        [16].12   // Node 3 message write error flag
        [0].12   // Node 2 Message Write Error Flag
        [32].12   // Node 4 message write error flag
        [48].12   // Node 5 message write error flag
        [64].12   // Node 6 message write error flag
        [16]   // Node 3 message write output data control block
        [80].12   // Node 7 message write error flag
        [96].12   // Node 8 message write error flag
        [2]   // FV2 Temperature Scaled -100/+400 tenths degree C
   FV_N101 : INT[255] := ([0] := 152, [1] := 60, [2] := 60, [3] := 586, [4] := 32767, [5] := 1107, [6] := 169, [7] := 117, [9] := 70, [10] := 110);   // FV INT Fermentation control integer workspace
        [9]   // Temp.register
        [7]   // Pointer to vessel's data file
        [35]   // Checkword Pointer
        [0]   // FV Data File Pointer
        [4]   // Next breakpoint time
        [1]   // Setpoint at previous breakpoint
        [30]   // PV550 Manual Valve Control Valve Checkword Number
        [2]   // Setpoint at next breakpoint
        [12]   // Operator Interface CT1 Manual Operation Value
        [14]   // Operator Interface CT2 Manual Operation Value
        [3]   // Previous breakpoint time
        [16]   // Operator Interface CT3 Manual Operation Value
        [18]   // Operator Interface CT4 Manual Operation Value
        [30].15   // Stops Invalid Pointer Error If No Valves Selected On Op. Int
        [20]   // Operator Interface CT5 Manual Operation Value
        [22]   // Operator Interface CT6 Manual Operation Value
        [38]   // Copy Of Current Checkword Manual Enabled Flag
        [32]   // Copy Of Current Checkword Energised Input Flag
        [37]   // Copy Of Current Checkword Energised Input Flag
        [36]   // Valve Operation 1 Open 2 Close 3 Auto
        [8]   // Fermenting Room PV550 data file pointer
        [6]   // Temporary result register
        [15].0   // Current Valve Manual/ Auto(PLC)
        [11].0   // Current Valve Energised/ De-energised
        [13].0   // Current Valve Energised/ De-energised
        [5]   // Time since last B.P in 1/10 hour
   FV_N104 : INT[255] := ([0] := -32768, [1] := -32768, [2] := -32768, [3] := -32768, [4] := -32768, [5] := -32768, [6] := -32768, [7] := -32768, [8] := -32768, [9] := -32768, [10] := -32768, [11] := -32768, [12] := -32768, [13] := -32768, [14] := -32768, [15] := -32768, [16] := -32768, [17] := -32768, [18] := -32768, [19] := -32768, [20] := -32768, [21] := -32768, [22] := -32768, [23] := -32768, [24] := -32768);   // FV_PC_BUF PC>PLC Fermentation Control Command Buff er File
        [23]   // PC>PLC FV System Command Buffer Command Type 1=Start,2=Stop 3=Modify Control
        [11]   // PC>PLC FV System Command Buffer Breakpoint F Time
        [13]   // PC>PLC FV System Command Buffer Breakpoint G Time
        [1]   // PC>PLC FV System Command Buffer Breakpoint A Time
        [3]   // PC>PLC FV System Command Buffer Breakpoint B Time
        [5]   // PC>PLC FV System Command Buffer Breakpoint C Time
        [7]   // PC>PLC FV System Command Buffer Breakpoint D Time
        [9]   // PC>PLC FV System Command Buffer Breakpoint E Time
        [2]   // PC>PLC FV System Command Buffer Breakpoint A Temperature Setpoint
        [4]   // PC>PLC FV System Command Buffer Breakpoint B Temperature Setpoint
        [6]   // PC>PLC FV System Command Buffer Breakpoint C Temperature Setpoint
        [8]   // PC>PLC FV System Command Buffer Breakpoint D Temperature Setpoint
        [0]   // PC>PLC FV System Vessel Number 1-28 = FV1-25,YSV1-3 95-96 YST1-2
        [15].4   // FV System PC Command Buffer Control Flags 1=Ageing Profile
        [15].6   // FV System PC Command Buffer Control Flags 1=Wait for yeast
        [10]   // PC>PLC FV System Command Buffer Breakpoint E Temperature Setpoint
        [12]   // PC>PLC FV System Command Buffer Breakpoint F Temperature Setpoint
        [14]   // PC>PLC FV System Command Buffer Breakpoint G Temperature Setpoint
        [15]   // PC>PLC FV System Command Buffer Profile Control / Configuration Flags
        [24]   // FV System PC Command Buffer Phase Number
        [16]   // PC>PLC FV System Command Buffer PC Private Flags
   FV_N11 : INT[255] := ([0] := 1, [32] := -1028);   // LOOP NO.
        [11].0   // Me>Node 5 heartbeat bit
        [14].0   // Me>Node 6 heartbeat bit
        [17].0   // Me>Node 7 heartbeat bit
        [20].0   // Me>Node 8 heartbeat bit
        [9].1   // BHP_RS Borehole Pump Start Signal Node 5 Output 1
        [2]   // Me>Node 2 Flags
        [0].0   // NODE 2 Outputs CT1 cooling valve drive flag
        [0]   // Check Loop Counter In Range
        [0].1   // NODE 2 Outputs CT2 cooling valve drive flag
        [11].1   // Node 5 to resend data
        [14].1   // Node 6 to resend data
        [0].6   // NODE 2 Outputs Fridge 1 Remote Start flag
        [0].2   // NODE 2 Outputs CT3 cooling valve drive flag
        [0].3   // NODE 2 Outputs CT4 cooling valve drive flag
        [170]   // Me>Node 7 heartbeat bit
        [17].1   // Node 7 to resend data
        [20].1   // Node 8 to resend data
        [2].0   // Me>Node 2 heartbeat bit
        [0].7   // NODE 2 Outputs Glycol recirc pump start flag
        [5].0   // Me>Node 3 heartbeat bit
        [0].4   // NODE 2 Outputs CT5 cooling valve drive flag
        [8].0   // Me>Node 4 heartbeat bit
        [0].5   // NODE 2 Outputs CT6 cooling valve drive flag
        [15]   // Move Binary Image Back To Node 7 Outputs
        [2].1   // Node 2 to resend data
        [5].1   // Node 3 to resend data
        [8].1   // Node 4 to resend data
   FV_N110 : INT[255] := ([0] := 231, [2] := 170, [3] := 100, [4] := 190, [5] := 275, [6] := 190, [7] := 305, [8] := 160, [9] := 486, [10] := 160, [11] := 586, [12] := 60, [13] := 32767, [14] := 60, [15] := 64, [17] := -32767, [18] := -32767, [19] := 1680, [20] := 13, [22] := 1693, [23] := 3, [24] := 6, [25] := 60, [26] := 60, [27] := 1693, [29] := 2, [30] := 24, [40] := 3, [41] := 59);   // FV DATA 0 CURRENT FV DATA
        [29]   // FLAGS - PLC CONTROL
        [28]   // CURRENT VOLUME HL*10
        [41]   // Cone ACTUAL TEMPERATURE -DEGREES 'C'*10
        [19]   // Current FV max. fermentation time
        [1]   // TEMPERATURE BREAKPOINT A. TIME 1/10 HOURS(ALWAYS=0)
        [29].1   // Current vessel deferred chilling enabled flag
        [3]   // TEMPERATURE BREAKPOINT B. TIME 1/10 HOURS(ALWAYS=0)
        [11]   // TEMPERATURE BREAKPOINT F. TIME 1/10 HOURS(ALWAYS=0)
        [13]   // TEMPERATURE BREAKPOINT G. TIME 1/10 HOURS(ALWAYS=0)
        [5]   // TEMPERATURE BREAKPOINT C. TIME 1/10 HOURS(ALWAYS=0)
        [7]   // TEMPERATURE BREAKPOINT D. TIME 1/10 HOURS(ALWAYS=0)
        [9]   // TEMPERATURE BREAKPOINT E. TIME 1/10 HOURS(ALWAYS=0)
        [30].5   // Current vessel deferred chilling temp.high flag
        [22]   // Current FV total residence time
        [15].5   // Profile Control Flags : This is a conditioning profile
        [15].3   // PLC TO USE CONE COOLING JACKET
        [15].9   // Current vessel deferred chilling manual override
        [20]   // Current FV warm conditioning time
        [27]   // CURRENT ELAPSED HOURS *10
        [40]   // FV Routing Status 9=Dirty
        [30].0   // Jacket Cooling Valve to open
        [26]   // Calculated Setpoint 1/10 degrees C
        [29].0   // PC TO SAVE TEMPERATURE DATA
        [15]   // FLAGS-PROFILE CONTROL
        [24]   // Phase0=No control 1to6 =Fermenting 8 =Pitching Hold 10 =Maturation 11to16=Conditioning
        [10]   // TEMPERATURE SETPOINT E. 1/10 DEGREE 'C'
        [15].2   // PLC TO FOLLOW RAMP Breakpoints A to B
        [12]   // TEMPERATURE SETPOINT F. 1/10 DEGREE 'C'
        [14]   // TEMPERATURE SETPOINT G. 1/10 DEGREE 'C'
        [36]   // Current vessel time to deferred chlling start (hrs.x10)
        [16].1   // Profile control flag Hold at B.P B
        [16].2   // Profile control flag Hold at B.P C
        [30].3   // Current vessel deferred chilling active
        [16].3   // Profile control flag Hold at B.P D
        [16].4   // Profile control flag Hold at B.P E
        [0]   // FV SYSTEM WORKING BUFFER VESSEL NUMBER
        [2]   // TEMPERATURE SETPOINT A. 1/10 DEGREE 'C'
        [16].5   // Profile control flag Hold at B.P F
        [16].6   // Profile control flag Hold at B.P G
        [30].4   // Current vessel final temp.reached
        [4]   // TEMPERATURE SETPOINT B. 1/10 DEGREE 'C'
        [6]   // TEMPERATURE SETPOINT C. 1/10 DEGREE 'C'
        [8]   // TEMPERATURE SETPOINT D. 1/10 DEGREE 'C'
        [30].1   // Cone Cooling Valve to open
        [25]   // Jacket ACTUAL TEMPERATURE -DEGREES 'C'*10
        [15].4   // Profile Control Flags : This is a maturation profile
   FV_N111 : INT[50] := ([0] := 1, [2] := 175, [3] := 200, [4] := 200, [5] := 440, [6] := 200, [7] := 480, [8] := 180, [9] := 650, [10] := 180, [11] := 820, [12] := 60, [13] := 32767, [14] := 60, [15] := 64, [16] := 20, [17] := -32767, [18] := -32767, [19] := 1680, [22] := 253, [23] := 1, [24] := 2, [25] := 199, [26] := 200, [27] := 253);   // FV1, CURRENT FV DATA
        [27]   // FV1,CURRENT ELAPSED HOURS *10
        [40]   // FV1,FV Routing Status 9=Dirty
        [36]   // FV1,Current vessel time to deferred chlling start (hrs.x10)
        [30].1   // FV1,Cone Cooling Valve to open
        [15].5   // FV1,Profile Control Flags : This is a conditioning profile
        [15]   // FV1,FLAGS-PROFILE CONTROL
        [30].3   // FV1,Current vessel deferred chilling active
        [24]   // FV1,Phase0=No control 1to6 =Fermenting 8 =Pitching Hold 10 =Maturation 11to16=Conditioning
        [15].4   // FV1,Profile Control Flags : This is a maturation profile
        [25]   // FV1,Jacket ACTUAL TEMPERATURE -DEGREES 'C'*10
        [15].2   // FV1,PLC TO FOLLOW RAMP Breakpoints A to B
        [29]   // FV1,FLAGS - PLC CONTROL
        [0]   // FV1,FV SYSTEM WORKING BUFFER VESSEL NUMBER
        [2]   // FV1,TEMPERATURE SETPOINT A. 1/10 DEGREE 'C'
        [30].4   // FV1,Current vessel final temp.reached
        [4]   // FV1,TEMPERATURE SETPOINT B. 1/10 DEGREE 'C'
        [6]   // FV1,TEMPERATURE SETPOINT C. 1/10 DEGREE 'C'
        [8]   // FV1,TEMPERATURE SETPOINT D. 1/10 DEGREE 'C'
        [11]   // FV1,TEMPERATURE BREAKPOINT F. TIME 1/10 HOURS(ALWAYS=0)
        [13]   // FV1,TEMPERATURE BREAKPOINT G. TIME 1/10 HOURS(ALWAYS=0)
        [30].5   // FV1,Current vessel deferred chilling temp.high flag
        [28]   // FV1,CURRENT VOLUME HL*10
        [15].3   // FV1,PLC TO USE CONE COOLING JACKET
        [41]   // FV1,Cone ACTUAL TEMPERATURE -DEGREES 'C'*10
        [26]   // FV1,Calculated Setpoint 1/10 degrees C
        [19]   // FV1,Current FV max. fermentation time
        [20]   // FV1,Current FV warm conditioning time
        [22]   // FV1,Current FV total residence time
        [29].0   // FV1,PC TO SAVE TEMPERATURE DATA
        [1]   // FV1,TEMPERATURE BREAKPOINT A. TIME 1/10 HOURS(ALWAYS=0)
        [29].1   // FV1,Current vessel deferred chilling enabled flag
        [30].0   // FV1,Jacket Cooling Valve to open
        [3]   // FV1,TEMPERATURE BREAKPOINT B. TIME 1/10 HOURS(ALWAYS=0)
        [5]   // FV1,TEMPERATURE BREAKPOINT C. TIME 1/10 HOURS(ALWAYS=0)
        [7]   // FV1,TEMPERATURE BREAKPOINT D. TIME 1/10 HOURS(ALWAYS=0)
        [9]   // FV1,TEMPERATURE BREAKPOINT E. TIME 1/10 HOURS(ALWAYS=0)
        [16].1   // FV1,Profile control flag Hold at B.P B
        [16].2   // FV1,Profile control flag Hold at B.P C
        [16].3   // FV1,Profile control flag Hold at B.P D
        [16].4   // FV1,Profile control flag Hold at B.P E
        [16].5   // FV1,Profile control flag Hold at B.P F
        [16].6   // FV1,Profile control flag Hold at B.P G
        [10]   // FV1,TEMPERATURE SETPOINT E. 1/10 DEGREE 'C'
        [15].9   // FV1,Current vessel deferred chilling manual override
        [12]   // FV1,TEMPERATURE SETPOINT F. 1/10 DEGREE 'C'
        [14]   // FV1,TEMPERATURE SETPOINT G. 1/10 DEGREE 'C'
   FV_N112 : INT[50] := ([0] := 2, [2] := 170, [3] := 100, [4] := 190, [5] := 264, [6] := 190, [7] := 290, [8] := 160, [9] := 532, [10] := 160, [11] := 632, [12] := 60, [13] := 32767, [14] := 60, [15] := 64, [17] := -32767, [18] := -32767, [19] := 1680, [20] := 15, [22] := 1695, [23] := 3, [24] := 6, [25] := 60, [26] := 60, [27] := 1695, [29] := 2, [30] := 24);   // FV2, CURRENT FV DATA
        [27]   // FV2,CURRENT ELAPSED HOURS *10
        [40]   // FV2,FV Routing Status 9=Dirty
        [36]   // FV2,Current vessel time to deferred chlling start (hrs.x10)
        [30].1   // FV2,Cone Cooling Valve to open
        [15]   // FV2,FLAGS-PROFILE CONTROL
        [15].5   // FV2,Profile Control Flags : This is a conditioning profile
        [30].3   // FV2,Current vessel deferred chilling active
        [24]   // FV2,Phase0=No control 1to6 =Fermenting 8 =Pitching Hold 10 =Maturation 11to16=Conditioning
        [15].4   // FV2,Profile Control Flags : This is a maturation profile
        [25]   // FV2,Jacket ACTUAL TEMPERATURE -DEGREES 'C'*10
        [15].2   // FV2,PLC TO FOLLOW RAMP Breakpoints A to B
        [29]   // FV2,FLAGS - PLC CONTROL
        [0]   // FV2,FV SYSTEM WORKING BUFFER VESSEL NUMBER
        [2]   // FV2,TEMPERATURE SETPOINT A. 1/10 DEGREE 'C'
        [30].4   // FV2,Current vessel final temp.reached
        [4]   // FV2,TEMPERATURE SETPOINT B. 1/10 DEGREE 'C'
        [6]   // FV2,TEMPERATURE SETPOINT C. 1/10 DEGREE 'C'
        [8]   // FV2,TEMPERATURE SETPOINT D. 1/10 DEGREE 'C'
        [11]   // FV2,TEMPERATURE BREAKPOINT F. TIME 1/10 HOURS(ALWAYS=0)
        [13]   // FV2,TEMPERATURE BREAKPOINT G. TIME 1/10 HOURS(ALWAYS=0)
        [15].3   // FV2,PLC TO USE CONE COOLING JACKET
        [30].5   // FV2,Current vessel deferred chilling temp.high flag
        [19]   // FV2,Current FV max. fermentation time
        [28]   // FV2,CURRENT VOLUME HL*10
        [41]   // FV2,Cone ACTUAL TEMPERATURE -DEGREES 'C'*10
        [26]   // FV2,Calculated Setpoint 1/10 degrees C
        [1]   // FV2,TEMPERATURE BREAKPOINT A. TIME 1/10 HOURS(ALWAYS=0)
        [29].1   // FV2,Current vessel deferred chilling enabled flag
        [20]   // FV2,Current FV warm conditioning time
        [3]   // FV2,TEMPERATURE BREAKPOINT B. TIME 1/10 HOURS(ALWAYS=0)
        [22]   // FV2,Current FV total residence time
        [29].0   // FV2,PC TO SAVE TEMPERATURE DATA
        [5]   // FV2,TEMPERATURE BREAKPOINT C. TIME 1/10 HOURS(ALWAYS=0)
        [7]   // FV2,TEMPERATURE BREAKPOINT D. TIME 1/10 HOURS(ALWAYS=0)
        [9]   // FV2,TEMPERATURE BREAKPOINT E. TIME 1/10 HOURS(ALWAYS=0)
        [30].0   // FV2,Jacket Cooling Valve to open
        [16].1   // FV2,Profile control flag Hold at B.P B
        [16].2   // FV2,Profile control flag Hold at B.P C
        [16].3   // FV2,Profile control flag Hold at B.P D
        [16].4   // FV2,Profile control flag Hold at B.P E
        [16].5   // FV2,Profile control flag Hold at B.P F
        [16].6   // FV2,Profile control flag Hold at B.P G
        [15].9   // FV2,Current vessel deferred chilling manual override
        [10]   // FV2,TEMPERATURE SETPOINT E. 1/10 DEGREE 'C'
        [12]   // FV2,TEMPERATURE SETPOINT F. 1/10 DEGREE 'C'
        [14]   // FV2,TEMPERATURE SETPOINT G. 1/10 DEGREE 'C'
   FV_N113 : INT[50] := ([0] := 3, [1] := -32767, [2] := -32767, [3] := -32767, [4] := -32767, [5] := -32767, [6] := -32767, [7] := -32767, [8] := -32767, [9] := -32767, [10] := -32767, [11] := -32767, [12] := -32767, [13] := -32767, [14] := -32767, [15] := -32767, [16] := -32767, [17] := -32767, [18] := -32767, [19] := -32767, [20] := -32767, [21] := -32767, [22] := -32767, [23] := 2, [25] := 431, [30] := 32);   // FV3, CURRENT FV DATA
        [27]   // FV3,CURRENT ELAPSED HOURS *10
        [40]   // FV3,FV Routing Status 9=Dirty
        [36]   // FV3,Current vessel time to deferred chlling start (hrs.x10)
        [30].1   // FV3,Cone Cooling Valve to open
        [15]   // FV3,FLAGS-PROFILE CONTROL
        [15].5   // FV3,Profile Control Flags : This is a conditioning profile
        [30].3   // FV3,Current vessel deferred chilling active
        [24]   // FV3,Phase0=No control 1to6 =Fermenting 8 =Pitching Hold 10 =Maturation 11to16=Conditioning
        [15].4   // FV3,Profile Control Flags : This is a maturation profile
        [25]   // FV3,Jacket ACTUAL TEMPERATURE -DEGREES 'C'*10
        [15].2   // FV3,PLC TO FOLLOW RAMP Breakpoints A to B
        [29]   // FV3,FLAGS - PLC CONTROL
        [0]   // FV3,FV SYSTEM WORKING BUFFER VESSEL NUMBER
        [2]   // FV3,TEMPERATURE SETPOINT A. 1/10 DEGREE 'C'
        [30].4   // FV3,Current vessel final temp.reached
        [4]   // FV3,TEMPERATURE SETPOINT B. 1/10 DEGREE 'C'
        [6]   // FV3,TEMPERATURE SETPOINT C. 1/10 DEGREE 'C'
        [8]   // FV3,TEMPERATURE SETPOINT D. 1/10 DEGREE 'C'
        [19]   // FV3,Current FV max. fermentation time
        [1]   // FV3,TEMPERATURE BREAKPOINT A. TIME 1/10 HOURS(ALWAYS=0)
        [20]   // FV3,Current FV warm conditioning time
        [29].1   // FV3,Current vessel deferred chilling enabled flag
        [3]   // FV3,TEMPERATURE BREAKPOINT B. TIME 1/10 HOURS(ALWAYS=0)
        [11]   // FV3,TEMPERATURE BREAKPOINT F. TIME 1/10 HOURS(ALWAYS=0)
        [13]   // FV3,TEMPERATURE BREAKPOINT G. TIME 1/10 HOURS(ALWAYS=0)
        [30].5   // FV3,Current vessel deferred chilling temp.high flag
        [28]   // FV3,CURRENT VOLUME HL*10
        [5]   // FV3,TEMPERATURE BREAKPOINT C. TIME 1/10 HOURS(ALWAYS=0)
        [15].3   // FV3,PLC TO USE CONE COOLING JACKET
        [26]   // FV3,Calculated Setpoint 1/10 degrees C
        [7]   // FV3,TEMPERATURE BREAKPOINT D. TIME 1/10 HOURS(ALWAYS=0)
        [41]   // FV3,Cone ACTUAL TEMPERATURE -DEGREES 'C'*10
        [9]   // FV3,TEMPERATURE BREAKPOINT E. TIME 1/10 HOURS(ALWAYS=0)
        [22]   // FV3,Current FV total residence time
        [29].0   // FV3,PC TO SAVE TEMPERATURE DATA
        [30].0   // FV3,Jacket Cooling Valve to open
        [16].1   // FV3,Profile control flag Hold at B.P B
        [16].2   // FV3,Profile control flag Hold at B.P C
        [16].3   // FV3,Profile control flag Hold at B.P D
        [10]   // FV3,TEMPERATURE SETPOINT E. 1/10 DEGREE 'C'
        [16].4   // FV3,Profile control flag Hold at B.P E
        [16].5   // FV3,Profile control flag Hold at B.P F
        [16].6   // FV3,Profile control flag Hold at B.P G
        [15].9   // FV3,Current vessel deferred chilling manual override
        [12]   // FV3,TEMPERATURE SETPOINT F. 1/10 DEGREE 'C'
        [14]   // FV3,TEMPERATURE SETPOINT G. 1/10 DEGREE 'C'
   FV_N114 : INT[50] := ([0] := 4, [2] := 240, [3] := 100, [4] := 240, [5] := 280, [6] := 240, [7] := 340, [8] := 240, [9] := 500, [10] := 240, [11] := 710, [12] := 240, [13] := 32767, [14] := 235, [17] := -32767, [18] := -32767, [19] := 14400, [20] := 18367, [22] := 32767, [23] := 3, [24] := 1, [25] := 247, [26] := 240, [27] := -9629, [29] := 2, [30] := 24);   // FV4, CURRENT FV DATA
        [15]   // FV4,FLAGS-PROFILE CONTROL
        [27]   // FV4,CURRENT ELAPSED HOURS *10
        [40]   // FV4,FV Routing Status 9=Dirty
        [36]   // FV4,Current vessel time to deferred chlling start (hrs.x10)
        [30].1   // FV4,Cone Cooling Valve to open
        [15].5   // FV4,Profile Control Flags : This is a conditioning profile
        [30].3   // FV4,Current vessel deferred chilling active
        [24]   // FV4,Phase0=No control 1to6 =Fermenting 8 =Pitching Hold 10 =Maturation 11to16=Conditioning
        [15].4   // FV4,Profile Control Flags : This is a maturation profile
        [25]   // FV4,Jacket ACTUAL TEMPERATURE -DEGREES 'C'*10
        [0]   // FV4,FV SYSTEM WORKING BUFFER VESSEL NUMBER
        [15].2   // FV4,PLC TO FOLLOW RAMP Breakpoints A to B
        [2]   // FV4,TEMPERATURE SETPOINT A. 1/10 DEGREE 'C'
        [30].4   // FV4,Current vessel final temp.reached
        [4]   // FV4,TEMPERATURE SETPOINT B. 1/10 DEGREE 'C'
        [29]   // FV4,FLAGS - PLC CONTROL
        [6]   // FV4,TEMPERATURE SETPOINT C. 1/10 DEGREE 'C'
        [8]   // FV4,TEMPERATURE SETPOINT D. 1/10 DEGREE 'C'
        [28]   // FV4,CURRENT VOLUME HL*10
        [1]   // FV4,TEMPERATURE BREAKPOINT A. TIME 1/10 HOURS(ALWAYS=0)
        [29].1   // FV4,Current vessel deferred chilling enabled flag
        [3]   // FV4,TEMPERATURE BREAKPOINT B. TIME 1/10 HOURS(ALWAYS=0)
        [5]   // FV4,TEMPERATURE BREAKPOINT C. TIME 1/10 HOURS(ALWAYS=0)
        [7]   // FV4,TEMPERATURE BREAKPOINT D. TIME 1/10 HOURS(ALWAYS=0)
        [19]   // FV4,Current FV max. fermentation time
        [9]   // FV4,TEMPERATURE BREAKPOINT E. TIME 1/10 HOURS(ALWAYS=0)
        [20]   // FV4,Current FV warm conditioning time
        [11]   // FV4,TEMPERATURE BREAKPOINT F. TIME 1/10 HOURS(ALWAYS=0)
        [13]   // FV4,TEMPERATURE BREAKPOINT G. TIME 1/10 HOURS(ALWAYS=0)
        [30].5   // FV4,Current vessel deferred chilling temp.high flag
        [15].3   // FV4,PLC TO USE CONE COOLING JACKET
        [26]   // FV4,Calculated Setpoint 1/10 degrees C
        [41]   // FV4,Cone ACTUAL TEMPERATURE -DEGREES 'C'*10
        [22]   // FV4,Current FV total residence time
        [29].0   // FV4,PC TO SAVE TEMPERATURE DATA
        [30].0   // FV4,Jacket Cooling Valve to open
        [16].1   // FV4,Profile control flag Hold at B.P B
        [16].2   // FV4,Profile control flag Hold at B.P C
        [16].3   // FV4,Profile control flag Hold at B.P D
        [16].4   // FV4,Profile control flag Hold at B.P E
        [16].5   // FV4,Profile control flag Hold at B.P F
        [16].6   // FV4,Profile control flag Hold at B.P G
        [10]   // FV4,TEMPERATURE SETPOINT E. 1/10 DEGREE 'C'
        [12]   // FV4,TEMPERATURE SETPOINT F. 1/10 DEGREE 'C'
        [14]   // FV4,TEMPERATURE SETPOINT G. 1/10 DEGREE 'C'
        [15].9   // FV4,Current vessel deferred chilling manual override
   FV_N115 : INT[50] := ([0] := 5, [1] := -32767, [2] := -32767, [3] := -32767, [4] := -32767, [5] := -32767, [6] := -32767, [7] := -32767, [8] := -32767, [9] := -32767, [10] := -32767, [11] := -32767, [12] := -32767, [13] := -32767, [14] := -32767, [15] := -32767, [16] := -32767, [17] := -32767, [18] := -32767, [19] := -32767, [20] := -32767, [21] := -32767, [22] := -32767, [23] := 2, [25] := 224, [30] := 32);   // FV5, CURRENT FV DATA
        [15]   // FV5,FLAGS-PROFILE CONTROL
        [27]   // FV5,CURRENT ELAPSED HOURS *10
        [40]   // FV5,FV Routing Status 9=Dirty
        [36]   // FV5,Current vessel time to deferred chlling start (hrs.x10)
        [30].1   // FV5,Cone Cooling Valve to open
        [15].5   // FV5,Profile Control Flags : This is a conditioning profile
        [24]   // FV5,Phase0=No control 1to6 =Fermenting 8 =Pitching Hold 10 =Maturation 11to16=Conditioning
        [30].3   // FV5,Current vessel deferred chilling active
        [15].4   // FV5,Profile Control Flags : This is a maturation profile
        [25]   // FV5,Jacket ACTUAL TEMPERATURE -DEGREES 'C'*10
        [0]   // FV5,FV SYSTEM WORKING BUFFER VESSEL NUMBER
        [2]   // FV5,TEMPERATURE SETPOINT A. 1/10 DEGREE 'C'
        [30].4   // FV5,Current vessel final temp.reached
        [4]   // FV5,TEMPERATURE SETPOINT B. 1/10 DEGREE 'C'
        [6]   // FV5,TEMPERATURE SETPOINT C. 1/10 DEGREE 'C'
        [8]   // FV5,TEMPERATURE SETPOINT D. 1/10 DEGREE 'C'
        [15].2   // FV5,PLC TO FOLLOW RAMP Breakpoints A to B
        [29]   // FV5,FLAGS - PLC CONTROL
        [28]   // FV5,CURRENT VOLUME HL*10
        [1]   // FV5,TEMPERATURE BREAKPOINT A. TIME 1/10 HOURS(ALWAYS=0)
        [29].1   // FV5,Current vessel deferred chilling enabled flag
        [3]   // FV5,TEMPERATURE BREAKPOINT B. TIME 1/10 HOURS(ALWAYS=0)
        [5]   // FV5,TEMPERATURE BREAKPOINT C. TIME 1/10 HOURS(ALWAYS=0)
        [7]   // FV5,TEMPERATURE BREAKPOINT D. TIME 1/10 HOURS(ALWAYS=0)
        [9]   // FV5,TEMPERATURE BREAKPOINT E. TIME 1/10 HOURS(ALWAYS=0)
        [19]   // FV5,Current FV max. fermentation time
        [22]   // FV5,Current FV total residence time
        [20]   // FV5,Current FV warm conditioning time
        [29].0   // FV5,PC TO SAVE TEMPERATURE DATA
        [11]   // FV5,TEMPERATURE BREAKPOINT F. TIME 1/10 HOURS(ALWAYS=0)
        [13]   // FV5,TEMPERATURE BREAKPOINT G. TIME 1/10 HOURS(ALWAYS=0)
        [30].5   // FV5,Current vessel deferred chilling temp.high flag
        [15].3   // FV5,PLC TO USE CONE COOLING JACKET
        [26]   // FV5,Calculated Setpoint 1/10 degrees C
        [41]   // FV5,Cone ACTUAL TEMPERATURE -DEGREES 'C'*10
        [30].0   // FV5,Jacket Cooling Valve to open
        [16].1   // FV5,Profile control flag Hold at B.P B
        [16].2   // FV5,Profile control flag Hold at B.P C
        [16].3   // FV5,Profile control flag Hold at B.P D
        [16].4   // FV5,Profile control flag Hold at B.P E
        [16].5   // FV5,Profile control flag Hold at B.P F
        [16].6   // FV5,Profile control flag Hold at B.P G
        [10]   // FV5,TEMPERATURE SETPOINT E. 1/10 DEGREE 'C'
        [12]   // FV5,TEMPERATURE SETPOINT F. 1/10 DEGREE 'C'
        [14]   // FV5,TEMPERATURE SETPOINT G. 1/10 DEGREE 'C'
        [15].9   // FV5,Current vessel deferred chilling manual override
   FV_N116 : INT[50] := ([0] := 6, [2] := 170, [3] := 100, [4] := 190, [5] := 270, [6] := 190, [7] := 300, [8] := 160, [9] := 530, [10] := 160, [11] := 630, [12] := 60, [13] := 32767, [14] := 60, [15] := 64, [16] := 20, [17] := -32767, [18] := -32767, [19] := 1680, [22] := 15, [23] := 1, [24] := 1, [25] := 176, [26] := 190, [27] := 15);   // FV6, CURRENT FV DATA
        [15]   // FV6,FLAGS-PROFILE CONTROL
        [27]   // FV6,CURRENT ELAPSED HOURS *10
        [40]   // FV6,FV Routing Status 9=Dirty
        [36]   // FV6,Current vessel time to deferred chlling start (hrs.x10)
        [30].1   // FV6,Cone Cooling Valve to open
        [15].5   // FV6,Profile Control Flags : This is a conditioning profile
        [24]   // FV6,Phase0=No control 1to6 =Fermenting 8 =Pitching Hold 10 =Maturation 11to16=Conditioning
        [30].3   // FV6,Current vessel deferred chilling active
        [15].4   // FV6,Profile Control Flags : This is a maturation profile
        [0]   // FV6,FV SYSTEM WORKING BUFFER VESSEL NUMBER
        [2]   // FV6,TEMPERATURE SETPOINT A. 1/10 DEGREE 'C'
        [30].4   // FV6,Current vessel final temp.reached
        [25]   // FV6,Jacket ACTUAL TEMPERATURE -DEGREES 'C'*10
        [4]   // FV6,TEMPERATURE SETPOINT B. 1/10 DEGREE 'C'
        [6]   // FV6,TEMPERATURE SETPOINT C. 1/10 DEGREE 'C'
        [8]   // FV6,TEMPERATURE SETPOINT D. 1/10 DEGREE 'C'
        [15].2   // FV6,PLC TO FOLLOW RAMP Breakpoints A to B
        [29]   // FV6,FLAGS - PLC CONTROL
        [28]   // FV6,CURRENT VOLUME HL*10
        [1]   // FV6,TEMPERATURE BREAKPOINT A. TIME 1/10 HOURS(ALWAYS=0)
        [29].1   // FV6,Current vessel deferred chilling enabled flag
        [22]   // FV6,Current FV total residence time
        [3]   // FV6,TEMPERATURE BREAKPOINT B. TIME 1/10 HOURS(ALWAYS=0)
        [5]   // FV6,TEMPERATURE BREAKPOINT C. TIME 1/10 HOURS(ALWAYS=0)
        [7]   // FV6,TEMPERATURE BREAKPOINT D. TIME 1/10 HOURS(ALWAYS=0)
        [9]   // FV6,TEMPERATURE BREAKPOINT E. TIME 1/10 HOURS(ALWAYS=0)
        [29].0   // FV6,PC TO SAVE TEMPERATURE DATA
        [19]   // FV6,Current FV max. fermentation time
        [20]   // FV6,Current FV warm conditioning time
        [11]   // FV6,TEMPERATURE BREAKPOINT F. TIME 1/10 HOURS(ALWAYS=0)
        [13]   // FV6,TEMPERATURE BREAKPOINT G. TIME 1/10 HOURS(ALWAYS=0)
        [30].5   // FV6,Current vessel deferred chilling temp.high flag
        [15].3   // FV6,PLC TO USE CONE COOLING JACKET
        [26]   // FV6,Calculated Setpoint 1/10 degrees C
        [41]   // FV6,Cone ACTUAL TEMPERATURE -DEGREES 'C'*10
        [30].0   // FV6,Jacket Cooling Valve to open
        [16].1   // FV6,Profile control flag Hold at B.P B
        [16].2   // FV6,Profile control flag Hold at B.P C
        [16].3   // FV6,Profile control flag Hold at B.P D
        [16].4   // FV6,Profile control flag Hold at B.P E
        [16].5   // FV6,Profile control flag Hold at B.P F
        [16].6   // FV6,Profile control flag Hold at B.P G
        [10]   // FV6,TEMPERATURE SETPOINT E. 1/10 DEGREE 'C'
        [12]   // FV6,TEMPERATURE SETPOINT F. 1/10 DEGREE 'C'
        [14]   // FV6,TEMPERATURE SETPOINT G. 1/10 DEGREE 'C'
        [15].9   // FV6,Current vessel deferred chilling manual override
   FV_N117 : INT[50] := ([0] := 7, [1] := -32767, [2] := -32767, [3] := -32767, [4] := -32767, [5] := -32767, [6] := -32767, [7] := -32767, [8] := -32767, [9] := -32767, [10] := -32767, [11] := -32767, [12] := -32767, [13] := -32767, [14] := -32767, [15] := -32767, [16] := -32767, [17] := -32767, [18] := -32767, [19] := -32767, [20] := -32767, [21] := -32767, [22] := -32767, [23] := 2, [25] := 64, [30] := 32);   // FV7, CURRENT FV DATA
        [15]   // FV7,FLAGS-PROFILE CONTROL
        [27]   // FV7,CURRENT ELAPSED HOURS *10
        [40]   // FV7,FV Routing Status 9=Dirty
        [36]   // FV7,Current vessel time to deferred chlling start (hrs.x10)
        [30].1   // FV7,Cone Cooling Valve to open
        [0]   // FV7,FV SYSTEM WORKING BUFFER VESSEL NUMBER
        [2]   // FV7,TEMPERATURE SETPOINT A. 1/10 DEGREE 'C'
        [24]   // FV7,Phase0=No control 1to6 =Fermenting 8 =Pitching Hold 10 =Maturation 11to16=Conditioning
        [30].4   // FV7,Current vessel final temp.reached
        [15].5   // FV7,Profile Control Flags : This is a conditioning profile
        [30].3   // FV7,Current vessel deferred chilling active
        [15].4   // FV7,Profile Control Flags : This is a maturation profile
        [4]   // FV7,TEMPERATURE SETPOINT B. 1/10 DEGREE 'C'
        [6]   // FV7,TEMPERATURE SETPOINT C. 1/10 DEGREE 'C'
        [8]   // FV7,TEMPERATURE SETPOINT D. 1/10 DEGREE 'C'
        [25]   // FV7,Jacket ACTUAL TEMPERATURE -DEGREES 'C'*10
        [15].2   // FV7,PLC TO FOLLOW RAMP Breakpoints A to B
        [29]   // FV7,FLAGS - PLC CONTROL
        [22]   // FV7,Current FV total residence time
        [1]   // FV7,TEMPERATURE BREAKPOINT A. TIME 1/10 HOURS(ALWAYS=0)
        [29].1   // FV7,Current vessel deferred chilling enabled flag
        [3]   // FV7,TEMPERATURE BREAKPOINT B. TIME 1/10 HOURS(ALWAYS=0)
        [28]   // FV7,CURRENT VOLUME HL*10
        [5]   // FV7,TEMPERATURE BREAKPOINT C. TIME 1/10 HOURS(ALWAYS=0)
        [7]   // FV7,TEMPERATURE BREAKPOINT D. TIME 1/10 HOURS(ALWAYS=0)
        [9]   // FV7,TEMPERATURE BREAKPOINT E. TIME 1/10 HOURS(ALWAYS=0)
        [29].0   // FV7,PC TO SAVE TEMPERATURE DATA
        [19]   // FV7,Current FV max. fermentation time
        [20]   // FV7,Current FV warm conditioning time
        [11]   // FV7,TEMPERATURE BREAKPOINT F. TIME 1/10 HOURS(ALWAYS=0)
        [13]   // FV7,TEMPERATURE BREAKPOINT G. TIME 1/10 HOURS(ALWAYS=0)
        [30].5   // FV7,Current vessel deferred chilling temp.high flag
        [15].3   // FV7,PLC TO USE CONE COOLING JACKET
        [26]   // FV7,Calculated Setpoint 1/10 degrees C
        [41]   // FV7,Cone ACTUAL TEMPERATURE -DEGREES 'C'*10
        [30].0   // FV7,Jacket Cooling Valve to open
        [16].1   // FV7,Profile control flag Hold at B.P B
        [16].2   // FV7,Profile control flag Hold at B.P C
        [16].3   // FV7,Profile control flag Hold at B.P D
        [16].4   // FV7,Profile control flag Hold at B.P E
        [16].5   // FV7,Profile control flag Hold at B.P F
        [16].6   // FV7,Profile control flag Hold at B.P G
        [15].9   // FV7,Current vessel deferred chilling manual override
        [10]   // FV7,TEMPERATURE SETPOINT E. 1/10 DEGREE 'C'
        [12]   // FV7,TEMPERATURE SETPOINT F. 1/10 DEGREE 'C'
        [14]   // FV7,TEMPERATURE SETPOINT G. 1/10 DEGREE 'C'
   FV_N118 : INT[50] := ([0] := 8, [1] := -32767, [2] := -32767, [3] := -32767, [4] := -32767, [5] := -32767, [6] := -32767, [7] := -32767, [8] := -32767, [9] := -32767, [10] := -32767, [11] := -32767, [12] := -32767, [13] := -32767, [14] := -32767, [15] := -32767, [16] := -32767, [17] := -32767, [18] := -32767, [19] := -32767, [20] := -32767, [21] := -32767, [22] := -32767, [23] := 2, [25] := 297, [30] := 32);   // FV8, CURRENT FV DATA
        [15]   // FV8,FLAGS-PROFILE CONTROL
        [27]   // FV8,CURRENT ELAPSED HOURS *10
        [40]   // FV8,FV Routing Status 9=Dirty
        [36]   // FV8,Current vessel time to deferred chlling start (hrs.x10)
        [30].1   // FV8,Cone Cooling Valve to open
        [0]   // FV8,FV SYSTEM WORKING BUFFER VESSEL NUMBER
        [2]   // FV8,TEMPERATURE SETPOINT A. 1/10 DEGREE 'C'
        [30].4   // FV8,Current vessel final temp.reached
        [4]   // FV8,TEMPERATURE SETPOINT B. 1/10 DEGREE 'C'
        [6]   // FV8,TEMPERATURE SETPOINT C. 1/10 DEGREE 'C'
        [8]   // FV8,TEMPERATURE SETPOINT D. 1/10 DEGREE 'C'
        [24]   // FV8,Phase0=No control 1to6 =Fermenting 8 =Pitching Hold 10 =Maturation 11to16=Conditioning
        [15].5   // FV8,Profile Control Flags : This is a conditioning profile
        [30].3   // FV8,Current vessel deferred chilling active
        [15].4   // FV8,Profile Control Flags : This is a maturation profile
        [25]   // FV8,Jacket ACTUAL TEMPERATURE -DEGREES 'C'*10
        [15].2   // FV8,PLC TO FOLLOW RAMP Breakpoints A to B
        [29]   // FV8,FLAGS - PLC CONTROL
        [22]   // FV8,Current FV total residence time
        [29].0   // FV8,PC TO SAVE TEMPERATURE DATA
        [19]   // FV8,Current FV max. fermentation time
        [1]   // FV8,TEMPERATURE BREAKPOINT A. TIME 1/10 HOURS(ALWAYS=0)
        [29].1   // FV8,Current vessel deferred chilling enabled flag
        [3]   // FV8,TEMPERATURE BREAKPOINT B. TIME 1/10 HOURS(ALWAYS=0)
        [5]   // FV8,TEMPERATURE BREAKPOINT C. TIME 1/10 HOURS(ALWAYS=0)
        [28]   // FV8,CURRENT VOLUME HL*10
        [7]   // FV8,TEMPERATURE BREAKPOINT D. TIME 1/10 HOURS(ALWAYS=0)
        [9]   // FV8,TEMPERATURE BREAKPOINT E. TIME 1/10 HOURS(ALWAYS=0)
        [20]   // FV8,Current FV warm conditioning time
        [11]   // FV8,TEMPERATURE BREAKPOINT F. TIME 1/10 HOURS(ALWAYS=0)
        [13]   // FV8,TEMPERATURE BREAKPOINT G. TIME 1/10 HOURS(ALWAYS=0)
        [15].3   // FV8,PLC TO USE CONE COOLING JACKET
        [30].5   // FV8,Current vessel deferred chilling temp.high flag
        [26]   // FV8,Calculated Setpoint 1/10 degrees C
        [41]   // FV8,Cone ACTUAL TEMPERATURE -DEGREES 'C'*10
        [30].0   // FV8,Jacket Cooling Valve to open
        [16].1   // FV8,Profile control flag Hold at B.P B
        [16].2   // FV8,Profile control flag Hold at B.P C
        [16].3   // FV8,Profile control flag Hold at B.P D
        [16].4   // FV8,Profile control flag Hold at B.P E
        [16].5   // FV8,Profile control flag Hold at B.P F
        [16].6   // FV8,Profile control flag Hold at B.P G
        [15].9   // FV8,Current vessel deferred chilling manual override
        [10]   // FV8,TEMPERATURE SETPOINT E. 1/10 DEGREE 'C'
        [12]   // FV8,TEMPERATURE SETPOINT F. 1/10 DEGREE 'C'
        [14]   // FV8,TEMPERATURE SETPOINT G. 1/10 DEGREE 'C'
   FV_N119 : INT[50] := ([0] := 9, [2] := 175, [3] := 200, [4] := 200, [5] := 440, [6] := 200, [7] := 480, [8] := 180, [9] := 650, [10] := 180, [11] := 820, [12] := 60, [13] := 32767, [14] := 60, [15] := 64, [16] := 20, [17] := -32767, [18] := -32767, [19] := 1680, [22] := 237, [23] := 1, [24] := 2, [25] := 199, [26] := 200, [27] := 237);   // FV9, CURRENT FV DATA
        [15]   // FV9,FLAGS-PROFILE CONTROL
        [27]   // FV9,CURRENT ELAPSED HOURS *10
        [40]   // FV9,FV Routing Status 9=Dirty
        [11]   // FV9,TEMPERATURE BREAKPOINT F. TIME 1/10 HOURS(ALWAYS=0)
        [36]   // FV9,Current vessel time to deferred chlling start (hrs.x10)
        [0]   // FV9,FV SYSTEM WORKING BUFFER VESSEL NUMBER
        [15].5   // FV9,Profile Control Flags : This is a conditioning profile
        [30].1   // FV9,Cone Cooling Valve to open
        [2]   // FV9,TEMPERATURE SETPOINT A. 1/10 DEGREE 'C'
        [30].4   // FV9,Current vessel final temp.reached
        [4]   // FV9,TEMPERATURE SETPOINT B. 1/10 DEGREE 'C'
        [6]   // FV9,TEMPERATURE SETPOINT C. 1/10 DEGREE 'C'
        [8]   // FV9,TEMPERATURE SETPOINT D. 1/10 DEGREE 'C'
        [24]   // FV9,Phase0=No control 1to6 =Fermenting 8 =Pitching Hold 10 =Maturation 11to16=Conditioning
        [15].4   // FV9,Profile Control Flags : This is a maturation profile
        [30].3   // FV9,Current vessel deferred chilling active
        [25]   // FV9,Jacket ACTUAL TEMPERATURE -DEGREES 'C'*10
        [29]   // FV9,FLAGS - PLC CONTROL
        [15].2   // FV9,PLC TO FOLLOW RAMP Breakpoints A to B
        [22]   // FV9,Current FV total residence time
        [29].0   // FV9,PC TO SAVE TEMPERATURE DATA
        [28]   // FV9,CURRENT VOLUME HL*10
        [1]   // FV9,TEMPERATURE BREAKPOINT A. TIME 1/10 HOURS(ALWAYS=0)
        [19]   // FV9,Current FV max. fermentation time
        [29].1   // FV9,Current vessel deferred chilling enabled flag
        [3]   // FV9,TEMPERATURE BREAKPOINT B. TIME 1/10 HOURS(ALWAYS=0)
        [5]   // FV9,TEMPERATURE BREAKPOINT C. TIME 1/10 HOURS(ALWAYS=0)
        [7]   // FV9,TEMPERATURE BREAKPOINT D. TIME 1/10 HOURS(ALWAYS=0)
        [20]   // FV9,Current FV warm conditioning time
        [9]   // FV9,TEMPERATURE BREAKPOINT E. TIME 1/10 HOURS(ALWAYS=0)
        [15].3   // FV9,PLC TO USE CONE COOLING JACKET
        [26]   // FV9,Calculated Setpoint 1/10 degrees C
        [13]   // FV9,TEMPERATURE BREAKPOINT G. TIME 1/10 HOURS(ALWAYS=0)
        [30].5   // FV9,Current vessel deferred chilling temp.high flag
        [41]   // FV9,Cone ACTUAL TEMPERATURE -DEGREES 'C'*10
        [30].0   // FV9,Jacket Cooling Valve to open
        [16].1   // FV9,Profile control flag Hold at B.P B
        [16].2   // FV9,Profile control flag Hold at B.P C
        [16].3   // FV9,Profile control flag Hold at B.P D
        [16].4   // FV9,Profile control flag Hold at B.P E
        [16].5   // FV9,Profile control flag Hold at B.P F
        [16].6   // FV9,Profile control flag Hold at B.P G
        [15].9   // FV9,Current vessel deferred chilling manual override
        [10]   // FV9,TEMPERATURE SETPOINT E. 1/10 DEGREE 'C'
        [12]   // FV9,TEMPERATURE SETPOINT F. 1/10 DEGREE 'C'
        [14]   // FV9,TEMPERATURE SETPOINT G. 1/10 DEGREE 'C'
   FV_N12 : INT[255] := ([1] := 950, [2] := 3500, [3] := 3200, [4] := 130, [5] := 5, [6] := 300, [7] := 3300, [8] := 3600, [10] := 120, [11] := 13, [12] := 16, [13] := 30, [14] := 20, [26] := 2019, [27] := 3, [28] := 4, [29] := 6, [31] := 29, [32] := 480, [33] := 480, [34] := 720, [35] := 7, [39] := 10, [40] := 5, [41] := 2);   // SYS_PARMS System Parameter Fil e
        [32]   // Deferred chilling on fermentation delay (hrs.x10)
        [34]   // Deferred chilling on conditioning delay (hrs.x10)
        [4]   // YSV emptying Max allowed volume gain in YSV. Litres
        [26]   // PC>PLC Settings Current Year
        [37]   // Deferred chilling off time hour
        [14]   // Seat clean on time reseeding main
        [38]   // Deferred chilling off time min.
        [0].0   // PLC>PC Settings Reload Request
        [12]   // Reseeding final water flush time
        [10]   // Reseeding rouser on time
        [13]   // Seat clean off time Reseeding main
        [33]   // Deferred chilling on maturation delay (hrs.x10)
        [0]   // PLC>PC System Settings Reload Required
        [6]   // YSV rouser on during storage timer setting
        [39]   // Deferred chilling fermentation temp. high value
        [1]   // YSV1 Filling alarm weight
        [2]   // YSV2 Filling alarm weight
        [11]   // Reseeding initial water displacement time
        [3]   // YSV3 Filling alarm weight
        [5]   // YSV Pitching Minimum allowed pitch rate Litres/Min
        [35]   // Deferred chilling on time hour
        [40]   // Deferred chilling maturation temp.high value
        [41]   // Deferred chilling conditioning temp. high value
        [36]   // Deferred chilling on time min.
        [7]   // YSV rouser off during storage timer setting
   FV_N120 : INT[50] := ([0] := 10, [1] := -32767, [2] := -32767, [3] := -32767, [4] := -32767, [5] := -32767, [6] := -32767, [7] := -32767, [8] := -32767, [9] := -32767, [10] := -32767, [11] := -32767, [12] := -32767, [13] := -32767, [14] := -32767, [15] := -32767, [16] := -32767, [17] := -32767, [18] := -32767, [19] := -32767, [20] := -32767, [21] := -32767, [22] := -32767, [23] := 2, [25] := 229, [30] := 32);   // FV10, CURRENT FV DATA
        [15].2   // FV10,PLC TO FOLLOW RAMP Breakpoints A to B
        [15]   // FV10,FLAGS-PROFILE CONTROL
        [41]   // FV10,Cone ACTUAL TEMPERATURE -DEGREES 'C'*10
        [28]   // FV10,CURRENT VOLUME HL*10
        [24]   // FV10,Phase0=No control 1to6 =Fermenting 8 =Pitching Hold 10 =Maturation 11to16=Conditioning
        [30].1   // FV10,Cone Cooling Valve to open
        [30].0   // FV10,Jacket Cooling Valve to open
        [29]   // FV10,FLAGS - PLC CONTROL
        [15].3   // FV10,PLC TO USE CONE COOLING JACKET
        [19]   // FV10,Current FV max. fermentation time
        [20]   // FV10,Current FV warm conditioning time
        [25]   // FV10,Jacket ACTUAL TEMPERATURE -DEGREES 'C'*10
        [26]   // FV10,Calculated Setpoint 1/10 degrees C
        [10]   // FV10,TEMPERATURE SETPOINT E. 1/10 DEGREE 'C'
        [12]   // FV10,TEMPERATURE SETPOINT F. 1/10 DEGREE 'C'
        [14]   // FV10,TEMPERATURE SETPOINT G. 1/10 DEGREE 'C'
        [0]   // FV10,FV SYSTEM WORKING BUFFER VESSEL NUMBER
        [2]   // FV10,TEMPERATURE SETPOINT A. 1/10 DEGREE 'C'
        [22]   // FV10,Current FV total residence time
        [30].4   // FV10,Current vessel final temp.reached
        [29].0   // FV10,PC TO SAVE TEMPERATURE DATA
        [4]   // FV10,TEMPERATURE SETPOINT B. 1/10 DEGREE 'C'
        [6]   // FV10,TEMPERATURE SETPOINT C. 1/10 DEGREE 'C'
        [8]   // FV10,TEMPERATURE SETPOINT D. 1/10 DEGREE 'C'
        [30].3   // FV10,Current vessel deferred chilling active
        [11]   // FV10,TEMPERATURE BREAKPOINT F. TIME 1/10 HOURS(ALWAYS=0)
        [13]   // FV10,TEMPERATURE BREAKPOINT G. TIME 1/10 HOURS(ALWAYS=0)
        [30].5   // FV10,Current vessel deferred chilling temp.high flag
        [27]   // FV10,CURRENT ELAPSED HOURS *10
        [40]   // FV10,FV Routing Status 9=Dirty
        [16].1   // FV10,Profile control flag Hold at B.P B
        [16].2   // FV10,Profile control flag Hold at B.P C
        [16].3   // FV10,Profile control flag Hold at B.P D
        [16].4   // FV10,Profile control flag Hold at B.P E
        [16].5   // FV10,Profile control flag Hold at B.P F
        [16].6   // FV10,Profile control flag Hold at B.P G
        [15].4   // FV10,Profile Control Flags : This is a maturation profile
        [36]   // FV10,Current vessel time to deferred chlling start (hrs.x10)
        [1]   // FV10,TEMPERATURE BREAKPOINT A. TIME 1/10 HOURS(ALWAYS=0)
        [29].1   // FV10,Current vessel deferred chilling enabled flag
        [3]   // FV10,TEMPERATURE BREAKPOINT B. TIME 1/10 HOURS(ALWAYS=0)
        [5]   // FV10,TEMPERATURE BREAKPOINT C. TIME 1/10 HOURS(ALWAYS=0)
        [7]   // FV10,TEMPERATURE BREAKPOINT D. TIME 1/10 HOURS(ALWAYS=0)
        [9]   // FV10,TEMPERATURE BREAKPOINT E. TIME 1/10 HOURS(ALWAYS=0)
        [15].5   // FV10,Profile Control Flags : This is a conditioning profile
        [15].9   // FV10,Current vessel deferred chilling manual override
   FV_N121 : INT[50] := ([0] := 11, [1] := -32767, [2] := -32767, [3] := -32767, [4] := -32767, [5] := -32767, [6] := -32767, [7] := -32767, [8] := -32767, [9] := -32767, [10] := -32767, [11] := -32767, [12] := -32767, [13] := -32767, [14] := -32767, [15] := -32767, [16] := -32767, [17] := -32767, [18] := -32767, [19] := -32767, [20] := -32767, [21] := -32767, [22] := -32767, [23] := 2, [25] := 205, [30] := 32, [41] := 442);   // FV11, CURRENT FV DATA
        [15].2   // FV11,PLC TO FOLLOW RAMP Breakpoints A to B
        [15]   // FV11,FLAGS-PROFILE CONTROL
        [41]   // FV11,Cone ACTUAL TEMPERATURE -DEGREES 'C'*10
        [28]   // FV11,CURRENT VOLUME HL*10
        [24]   // FV11,Phase0=No control 1to6 =Fermenting 8 =Pitching Hold 10 =Maturation 11to16=Conditioning
        [30].1   // FV11,Cone Cooling Valve to open
        [30].0   // FV11,Jacket Cooling Valve to open
        [19]   // FV11,Current FV max. fermentation time
        [15].3   // FV11,PLC TO USE CONE COOLING JACKET
        [26]   // FV11,Calculated Setpoint 1/10 degrees C
        [29]   // FV11,FLAGS - PLC CONTROL
        [20]   // FV11,Current FV warm conditioning time
        [25]   // FV11,Jacket ACTUAL TEMPERATURE -DEGREES 'C'*10
        [10]   // FV11,TEMPERATURE SETPOINT E. 1/10 DEGREE 'C'
        [12]   // FV11,TEMPERATURE SETPOINT F. 1/10 DEGREE 'C'
        [14]   // FV11,TEMPERATURE SETPOINT G. 1/10 DEGREE 'C'
        [0]   // FV11,FV SYSTEM WORKING BUFFER VESSEL NUMBER
        [2]   // FV11,TEMPERATURE SETPOINT A. 1/10 DEGREE 'C'
        [30].4   // FV11,Current vessel final temp.reached
        [4]   // FV11,TEMPERATURE SETPOINT B. 1/10 DEGREE 'C'
        [22]   // FV11,Current FV total residence time
        [29].0   // FV11,PC TO SAVE TEMPERATURE DATA
        [6]   // FV11,TEMPERATURE SETPOINT C. 1/10 DEGREE 'C'
        [8]   // FV11,TEMPERATURE SETPOINT D. 1/10 DEGREE 'C'
        [30].3   // FV11,Current vessel deferred chilling active
        [11]   // FV11,TEMPERATURE BREAKPOINT F. TIME 1/10 HOURS(ALWAYS=0)
        [13]   // FV11,TEMPERATURE BREAKPOINT G. TIME 1/10 HOURS(ALWAYS=0)
        [30].5   // FV11,Current vessel deferred chilling temp.high flag
        [27]   // FV11,CURRENT ELAPSED HOURS *10
        [16].1   // FV11,Profile control flag Hold at B.P B
        [40]   // FV11,FV Routing Status 9=Dirty
        [16].2   // FV11,Profile control flag Hold at B.P C
        [16].3   // FV11,Profile control flag Hold at B.P D
        [16].4   // FV11,Profile control flag Hold at B.P E
        [16].5   // FV11,Profile control flag Hold at B.P F
        [16].6   // FV11,Profile control flag Hold at B.P G
        [15].4   // FV11,Profile Control Flags : This is a maturation profile
        [36]   // FV11,Current vessel time to deferred chlling start (hrs.x10)
        [1]   // FV11,TEMPERATURE BREAKPOINT A. TIME 1/10 HOURS(ALWAYS=0)
        [29].1   // FV11,Current vessel deferred chilling enabled flag
        [3]   // FV11,TEMPERATURE BREAKPOINT B. TIME 1/10 HOURS(ALWAYS=0)
        [5]   // FV11,TEMPERATURE BREAKPOINT C. TIME 1/10 HOURS(ALWAYS=0)
        [15].5   // FV11,Profile Control Flags : This is a conditioning profile
        [7]   // FV11,TEMPERATURE BREAKPOINT D. TIME 1/10 HOURS(ALWAYS=0)
        [9]   // FV11,TEMPERATURE BREAKPOINT E. TIME 1/10 HOURS(ALWAYS=0)
        [15].9   // FV11,Current vessel deferred chilling manual override
   FV_N122 : INT[50] := ([0] := 12, [2] := 170, [3] := 100, [4] := 190, [5] := 260, [6] := 190, [7] := 280, [8] := 160, [9] := 488, [10] := 160, [11] := 588, [12] := 60, [13] := 32767, [14] := 60, [15] := 64, [17] := -32767, [18] := -32767, [19] := 1680, [22] := 494, [23] := 3, [24] := 5, [25] := 154, [26] := 154, [27] := 494, [30] := 1);   // FV12, CURRENT FV DATA
        [15].2   // FV12,PLC TO FOLLOW RAMP Breakpoints A to B
        [15]   // FV12,FLAGS-PROFILE CONTROL
        [41]   // FV12,Cone ACTUAL TEMPERATURE -DEGREES 'C'*10
        [28]   // FV12,CURRENT VOLUME HL*10
        [24]   // FV12,Phase0=No control 1to6 =Fermenting 8 =Pitching Hold 10 =Maturation 11to16=Conditioning
        [30].1   // FV12,Cone Cooling Valve to open
        [15].3   // FV12,PLC TO USE CONE COOLING JACKET
        [25]   // FV12,Jacket ACTUAL TEMPERATURE -DEGREES 'C'*10
        [19]   // FV12,Current FV max. fermentation time
        [30].0   // FV12,Jacket Cooling Valve to open
        [26]   // FV12,Calculated Setpoint 1/10 degrees C
        [20]   // FV12,Current FV warm conditioning time
        [29]   // FV12,FLAGS - PLC CONTROL
        [10]   // FV12,TEMPERATURE SETPOINT E. 1/10 DEGREE 'C'
        [12]   // FV12,TEMPERATURE SETPOINT F. 1/10 DEGREE 'C'
        [14]   // FV12,TEMPERATURE SETPOINT G. 1/10 DEGREE 'C'
        [0]   // FV12,FV SYSTEM WORKING BUFFER VESSEL NUMBER
        [2]   // FV12,TEMPERATURE SETPOINT A. 1/10 DEGREE 'C'
        [30].4   // FV12,Current vessel final temp.reached
        [4]   // FV12,TEMPERATURE SETPOINT B. 1/10 DEGREE 'C'
        [6]   // FV12,TEMPERATURE SETPOINT C. 1/10 DEGREE 'C'
        [8]   // FV12,TEMPERATURE SETPOINT D. 1/10 DEGREE 'C'
        [22]   // FV12,Current FV total residence time
        [29].0   // FV12,PC TO SAVE TEMPERATURE DATA
        [30].3   // FV12,Current vessel deferred chilling active
        [11]   // FV12,TEMPERATURE BREAKPOINT F. TIME 1/10 HOURS(ALWAYS=0)
        [13]   // FV12,TEMPERATURE BREAKPOINT G. TIME 1/10 HOURS(ALWAYS=0)
        [30].5   // FV12,Current vessel deferred chilling temp.high flag
        [16].1   // FV12,Profile control flag Hold at B.P B
        [16].2   // FV12,Profile control flag Hold at B.P C
        [16].3   // FV12,Profile control flag Hold at B.P D
        [16].4   // FV12,Profile control flag Hold at B.P E
        [16].5   // FV12,Profile control flag Hold at B.P F
        [27]   // FV12,CURRENT ELAPSED HOURS *10
        [15].4   // FV12,Profile Control Flags : This is a maturation profile
        [40]   // FV12,FV Routing Status 9=Dirty
        [16].6   // FV12,Profile control flag Hold at B.P G
        [36]   // FV12,Current vessel time to deferred chlling start (hrs.x10)
